// TIA Portal project "V1.0Final" (V17)

(* hardware
DEVICE "S7-1200 station_1"  S7-1200 Station
   slot 0: "Rack_0"  S7-1200 Rack  Rack  V1.0
   slot 1: "PLC_1"  CPU 1212C AC/DC/Rly  6ES7 212-1BD30-0XB0  V2.0
   slot 2: "AI 4x13BIT_1"  6ES7 231-4HD32-0XB0  V2.1
   slot 3: "AQ 2x14BIT_1"  SM 1232 AQ2  6ES7 232-4HB32-0XB0  V2.1
DEVICE "HMI_1"  KTP700 Basic PN
   slot 0: "HMI_1"  KTP700 Basic PN  6AV2 123-2GB03-0AX0  17.0.0.0
   slot 1: "HMI_RT_1"  KTP700 Basic PN  6AV2 123-2GB03-0AX0  17.0.0.0
   slot 5: "HMI_1.IE_CP_1"  PROFINET Interface  17.0.0.0
      slot 1: "PROFINET Interface_1"  PROFINET Interface
         slot 1: "Port_1"  Port
*)

// ===== PLC "PLC_1"  CPU 1212C AC/DC/Rly =====

VAR_GLOBAL   // PLC tag table "Default tag table"
   "DI_EM_STOP" AT %I0.0 : Bool;
   "DI_LS_Tørrkjøringsvern" AT %I0.1 : Bool;
   "DI_Reset_EM_STOP" AT %I0.2 : Bool;
   "AI_LT_01" AT %IW100 : Int;
   "DQ_Lys_EM_STOP" AT %Q0.1 : Bool;
   "AQ1_PÅDRAG_PUMPE_01" AT %QW112 : Int;
   "AQ2" AT %QW114 : Int;
   "DI_PUMPE_01_KJØRER" AT %I0.3 : Bool;
   "Tag_1" AT %M0.0 : Bool;
   "DQ_START_PUMPE_01" AT %Q0.2 : Bool;
   "AI_Hastighet_P01" AT %IW102 : Int;
END_VAR

// folder: Equipment

TYPE "UDT_Analog_Konvertering"
   STRUCT
      CFG : Struct   // Configuration Data
         Spare : Bool;
      END_STRUCT;
      Sts : Struct   // Status Data
         EU_Verdi_Out : Real;
      END_STRUCT;
      Cmd : Struct   // Command and request Data
         Spare : Bool;
      END_STRUCT;
      Par : Struct   // Parameter Data
         EU_Min : Real;
         EU_Max : Real;
      END_STRUCT;
      Fit : Struct   // Warning and alarm triggers
         Feil : Bool;
      END_STRUCT;
      Spare : Bool;   // False
   END_STRUCT;
END_TYPE

TYPE "UDT_Pumpe_Kontroll"
   STRUCT
      CFG : Struct
         Spare : Bool;
      END_STRUCT;
      Sts : Struct
         Pumpe_Run : Bool;
         Pumpe_Status : Int;
         Pumpe_Faktisk_Hastighet_Fra_VFD : Real;
         Pumpe_Pådrag_Fra_PID_Blokk : Real;
      END_STRUCT;
      Cmd : Struct
         Man_Start_Pumpe : Bool;
         Man_Stop_Pumpe : Bool;
         Auto_Start_Pumpe : Bool;
         EM_Stop : Bool;
         Tørrkjøringsvakt_LS_01 : Bool;
      END_STRUCT;
      Par : Struct
         Pådrag_Fra_PID_Blokk : Int;
      END_STRUCT;
      Fit : Struct
         Feil : Bool;
      END_STRUCT;
   END_STRUCT;
END_TYPE

// folder: Machine

TYPE "UDT_HMI"
   STRUCT
      CFG : Struct
         Spare : Bool;
      END_STRUCT;
      Sts : Struct
         HMI_PV : Real;
         HMI_Pump_Status : Int;
      END_STRUCT;
      Cmd : Struct
         HMI_Pump_Auto : Bool;
         HMI_Pump_Manuell : Bool;
         HMI_Pump_Start : Bool;
         HMI_Pump_Stop : Bool;
         HMI_Reset_Alarm : Bool;
         Spare : Bool;
      END_STRUCT;
      Par : Struct
         HMI_P_Gain : Real;
         HMI_Ti : Real;
         HMI_Td : Real;
         HMI_Manual_Speed_Ref : Real;
         HMI_LT_Level_SP : Real;
         HMI_LT_EU_Min : Real;
         HMI_LT_EU_Max : Real;
         HMI_Anti_Windup : Bool;
         Spare : Bool;
      END_STRUCT;
      Fit : Struct
         HMI_EM_Stop_Alarm : Bool;
         HMI_LS_Activated : Bool;
         HMI_Fault_Timer_SP : Time;
         HMI_Fault : Bool;
      END_STRUCT;
   END_STRUCT;
END_TYPE

// folder: (top level)

DATA_BLOCK "LT_01"   // DB6
{ S7_Optimized_Access := 'TRUE' }
VERSION : 0.1
// stored: InstanceOfName Analog_Konvertering
"Analog_Konvertering"
BEGIN
END_DATA_BLOCK

DATA_BLOCK "Pumpe_01_Kontroll_DB"   // DB8
{ S7_Optimized_Access := 'TRUE' }
VERSION : 0.1
// stored: InstanceOfName Pumpe_Kontroll
"Pumpe_Kontroll"
BEGIN
END_DATA_BLOCK

DATA_BLOCK "Regulerings_Rig_01_DB"   // DB9
{ S7_Optimized_Access := 'TRUE' }
VERSION : 0.1
// stored: InstanceOfName Regulerings_Rig
"Regulerings_Rig"
BEGIN
END_DATA_BLOCK

DATA_BLOCK "VFD_AQ_Hastighet_Pumpe01_DB"   // DB11
{ S7_Optimized_Access := 'TRUE' }
VERSION : 0.1
// stored: InstanceOfName Analog_Konvertering
"Analog_Konvertering"
BEGIN
END_DATA_BLOCK

// folder: Global_Data

DATA_BLOCK "DB_Equipment"   // DB3
{ S7_Optimized_Access := 'TRUE' }
VERSION : 0.1
   VAR
      Pumpe_01_Kontroll : "UDT_Pumpe_Kontroll";
   END_VAR
   VAR RETAIN
      LT_01_Kontrolll : "UDT_Analog_Konvertering";
      HMI_Kontroll_Pumpe_01 : "UDT_HMI";
   END_VAR
   VAR
      VFD_01_Speed : "UDT_Analog_Konvertering";
   END_VAR
BEGIN
END_DATA_BLOCK

DATA_BLOCK "DB_Machine"   // DB4
{ S7_Optimized_Access := 'TRUE' }
VERSION : 0.1
   VAR
      HMI_Control : "UDT_HMI";
   END_VAR
BEGIN
END_DATA_BLOCK

// folder: System blocks/Program resources

DATA_BLOCK "EM_Stop_TON_DB"   // DB1
{ S7_Optimized_Access := 'TRUE' }
AUTHOR : Simatic
FAMILY : IEC
NAME : IEC_TMR
VERSION : 1.0
// stored: InstanceOfName IEC_TIMER
"IEC_TIMER"
BEGIN
END_DATA_BLOCK

DATA_BLOCK "EM_Stop_TOF_DB"   // DB2
{ S7_Optimized_Access := 'TRUE' }
AUTHOR : Simatic
FAMILY : IEC
NAME : IEC_TMR
VERSION : 1.0
// stored: InstanceOfName IEC_TIMER
"IEC_TIMER"
BEGIN
END_DATA_BLOCK

DATA_BLOCK "Pump_Fault_Timer_DB"   // DB5
{ S7_Optimized_Access := 'TRUE' }
AUTHOR : Simatic
FAMILY : IEC
NAME : IEC_TMR
VERSION : 1.0
// stored: InstanceOfName IEC_TIMER
"IEC_TIMER"
BEGIN
END_DATA_BLOCK

// folder: (top level)

ORGANIZATION_BLOCK "Main"   // OB1, LAD, ProgramCycle
TITLE = "Main Program Sweep (Cycle)"
{ S7_Optimized_Access := 'TRUE' }
VERSION : 0.1
BEGIN
END_ORGANIZATION_BLOCK

ORGANIZATION_BLOCK "Cyclic interrupt"   // OB30, LAD, CyclicInterrupt
{ S7_Optimized_Access := 'TRUE' }
VERSION : 0.1
   VAR_TEMP
      "0" : Bool;
   END_VAR
BEGIN

REGION Network 1
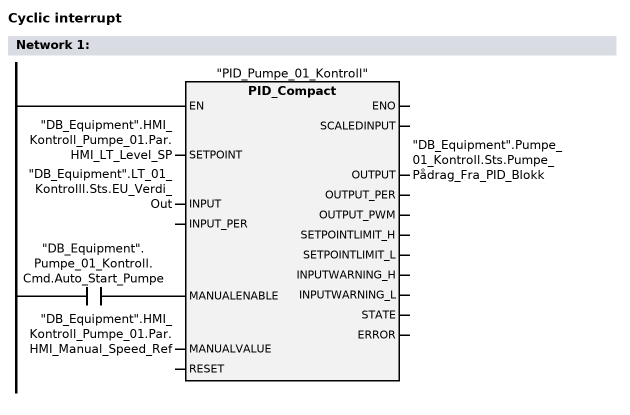
   "PID_Pumpe_01_Kontroll"(Setpoint := "DB_Equipment".HMI_Kontroll_Pumpe_01.Par.HMI_LT_Level_SP,   // PID_Compact
                           Input := "DB_Equipment".LT_01_Kontrolll.Sts.EU_Verdi_Out,
                           ManualEnable := "DB_Equipment".Pumpe_01_Kontroll.Cmd.Auto_Start_Pumpe,
                           ManualValue := "DB_Equipment".HMI_Kontroll_Pumpe_01.Par.HMI_Manual_Speed_Ref,
                           Output => "DB_Equipment".Pumpe_01_Kontroll.Sts.Pumpe_Pådrag_Fra_PID_Blokk);
END_REGION
END_ORGANIZATION_BLOCK

ORGANIZATION_BLOCK "Machine"   // OB123, LAD, ProgramCycle
TITLE = "Main Program Sweep (Cycle)"
{ S7_Optimized_Access := 'TRUE' }
VERSION : 0.1
BEGIN

REGION Network 1
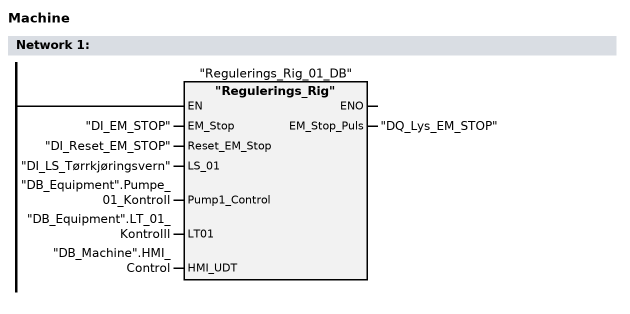
   RUNG wire#powerrail
      "Regulerings_Rig_01_DB"(EM_Stop := "DI_EM_STOP", Reset_EM_Stop := "DI_Reset_EM_STOP", LS_01 := "DI_LS_Tørrkjøringsvern", Pump1_Control := "DB_Equipment".Pumpe_01_Kontroll, LT01 := "DB_Equipment".LT_01_Kontrolll, HMI_UDT := "DB_Machine".HMI_Control, EM_Stop_Puls => "DQ_Lys_EM_STOP")
   END_RUNG
   // the same network as SCL:
   "Regulerings_Rig_01_DB"(EM_Stop := "DI_EM_STOP",   // "Regulerings_Rig"
                           Reset_EM_Stop := "DI_Reset_EM_STOP",
                           LS_01 := "DI_LS_Tørrkjøringsvern",
                           Pump1_Control := "DB_Equipment".Pumpe_01_Kontroll,
                           LT01 := "DB_Equipment".LT_01_Kontrolll,
                           HMI_UDT := "DB_Machine".HMI_Control,
                           EM_Stop_Puls => "DQ_Lys_EM_STOP");
END_REGION
END_ORGANIZATION_BLOCK

ORGANIZATION_BLOCK "Equipment"   // OB124, LAD, ProgramCycle
TITLE = "Main Program Sweep (Cycle)"
{ S7_Optimized_Access := 'TRUE' }
VERSION : 0.1
BEGIN

REGION Network 1
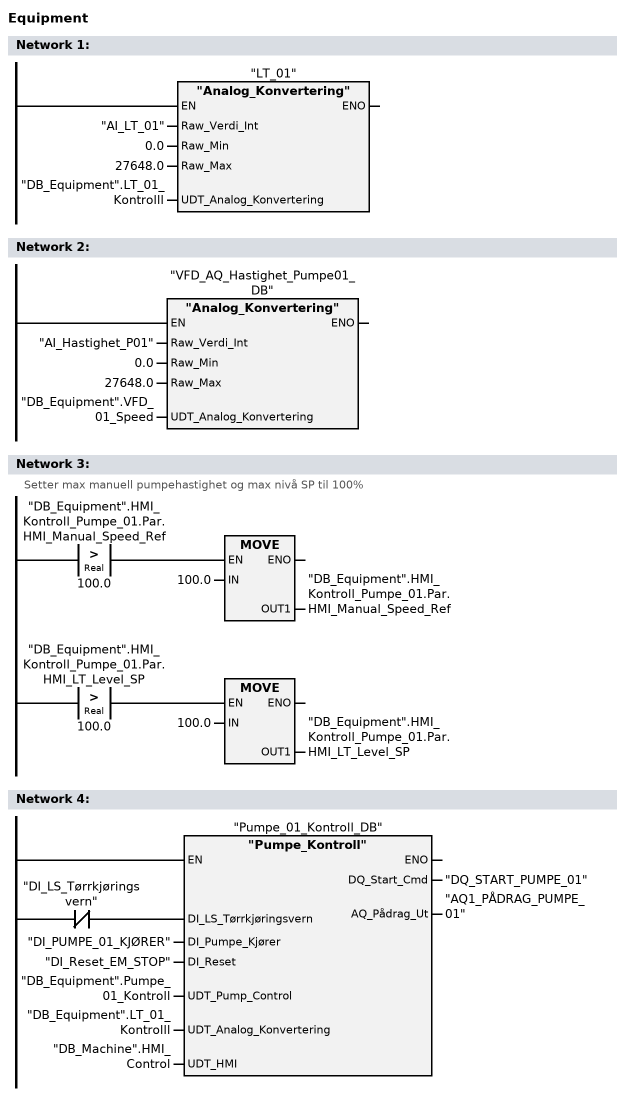
   RUNG wire#powerrail
      "LT_01"(Raw_Verdi_Int := "AI_LT_01", Raw_Min := 0.0, Raw_Max := 27648.0, UDT_Analog_Konvertering := "DB_Equipment".LT_01_Kontrolll)
   END_RUNG
   // the same network as SCL:
   "LT_01"(Raw_Verdi_Int := "AI_LT_01",   // "Analog_Konvertering"
           Raw_Min := 0.0,
           Raw_Max := 27648.0,
           UDT_Analog_Konvertering := "DB_Equipment".LT_01_Kontrolll);
END_REGION

REGION Network 2
   RUNG wire#powerrail
      "VFD_AQ_Hastighet_Pumpe01_DB"(Raw_Verdi_Int := "AI_Hastighet_P01", Raw_Min := 0.0, Raw_Max := 27648.0, UDT_Analog_Konvertering := "DB_Equipment".VFD_01_Speed)
   END_RUNG
   // the same network as SCL:
   "VFD_AQ_Hastighet_Pumpe01_DB"(Raw_Verdi_Int := "AI_Hastighet_P01",   // "Analog_Konvertering"
                           Raw_Min := 0.0,
                           Raw_Max := 27648.0,
                           UDT_Analog_Konvertering := "DB_Equipment".VFD_01_Speed);
END_REGION

REGION Network 3
   // Setter max manuell pumpehastighet og max nivå SP til 100%
   RUNG wire#powerrail
      { S7_Templates := "SrcType := Real" } GT_Contact(in1 := "DB_Equipment".HMI_Kontroll_Pumpe_01.Par.HMI_Manual_Speed_Ref, in2 := 100.0)
      { S7_GenerateENO := "TRUE" } Move(in := 100.0, out1 => "DB_Equipment".HMI_Kontroll_Pumpe_01.Par.HMI_Manual_Speed_Ref)
   END_RUNG
   RUNG wire#powerrail
      { S7_Templates := "SrcType := Real" } GT_Contact(in1 := "DB_Equipment".HMI_Kontroll_Pumpe_01.Par.HMI_LT_Level_SP, in2 := 100.0)
      { S7_GenerateENO := "TRUE" } Move(in := 100.0, out1 => "DB_Equipment".HMI_Kontroll_Pumpe_01.Par.HMI_LT_Level_SP)
   END_RUNG
   // the same network as SCL:
   IF "DB_Equipment".HMI_Kontroll_Pumpe_01.Par.HMI_Manual_Speed_Ref > 100.0 THEN
       "DB_Equipment".HMI_Kontroll_Pumpe_01.Par.HMI_Manual_Speed_Ref := 100.0;
   END_IF;
   IF "DB_Equipment".HMI_Kontroll_Pumpe_01.Par.HMI_LT_Level_SP > 100.0 THEN
       "DB_Equipment".HMI_Kontroll_Pumpe_01.Par.HMI_LT_Level_SP := 100.0;
   END_IF;
END_REGION

REGION Network 4
   RUNG wire#powerrail
      "Pumpe_01_Kontroll_DB"(DI_LS_Tørrkjøringsvern := wire#w1, DI_Pumpe_Kjører := "DI_PUMPE_01_KJØRER", DI_Reset := "DI_Reset_EM_STOP", UDT_Pump_Control := "DB_Equipment".Pumpe_01_Kontroll, UDT_Analog_Konvertering := "DB_Equipment".LT_01_Kontrolll, UDT_HMI := "DB_Machine".HMI_Control, DQ_Start_Cmd => "DQ_START_PUMPE_01", AQ_Pådrag_Ut => "AQ1_PÅDRAG_PUMPE_01")
   END_RUNG
   RUNG wire#powerrail
      I_Contact( "DI_LS_Tørrkjøringsvern" )
   END_RUNG wire#w1
   // the same network as SCL:
   "Pumpe_01_Kontroll_DB"(DI_LS_Tørrkjøringsvern := NOT "DI_LS_Tørrkjøringsvern",   // "Pumpe_Kontroll"
                          DI_Pumpe_Kjører := "DI_PUMPE_01_KJØRER",
                          DI_Reset := "DI_Reset_EM_STOP",
                          UDT_Pump_Control := "DB_Equipment".Pumpe_01_Kontroll,
                          UDT_Analog_Konvertering := "DB_Equipment".LT_01_Kontrolll,
                          UDT_HMI := "DB_Machine".HMI_Control,
                          DQ_Start_Cmd => "DQ_START_PUMPE_01",
                          AQ_Pådrag_Ut => "AQ1_PÅDRAG_PUMPE_01");
END_REGION
END_ORGANIZATION_BLOCK

// folder: Equipment

FUNCTION_BLOCK "Analog_Konvertering"   // FB2, LAD
{ S7_Optimized_Access := 'TRUE' }
VERSION : 0.1
   VAR_INPUT
      Raw_Verdi_Int : Int;
      Raw_Min : Real;
      Raw_Max : Real;
   END_VAR
   VAR_IN_OUT
      UDT_Analog_Konvertering : "UDT_Analog_Konvertering";
   END_VAR
   VAR
      Convert_Value : Real;
      Raw_Value_Real : Real;
      EU_Value_Real : Real;
   END_VAR
BEGIN

REGION Network 1
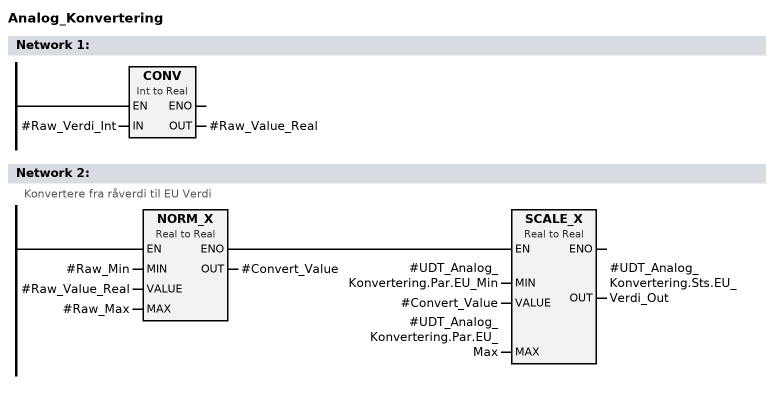
   RUNG wire#powerrail
      { S7_Templates := "[SrcType := Int, DestType := Real]"; S7_GenerateENO := "TRUE" } Convert(in := #Raw_Verdi_Int, out => #Raw_Value_Real)
   END_RUNG
   // the same network as SCL:
   #Raw_Value_Real := INT_TO_REAL(#Raw_Verdi_Int);
END_REGION

REGION Network 2
   // Konvertere fra råverdi til EU Verdi
   RUNG wire#powerrail
      { S7_Templates := "[SrcType := Real, DestType := Real]"; S7_GenerateENO := "TRUE" } Normalize(min := #Raw_Min, value := #Raw_Value_Real, max := #Raw_Max, out => #Convert_Value)
      { S7_Templates := "[SrcType := Real, DestType := Real]"; S7_GenerateENO := "TRUE" } Scale(min := #UDT_Analog_Konvertering.Par.EU_Min, value := #Convert_Value, max := #UDT_Analog_Konvertering.Par.EU_Max, out => #UDT_Analog_Konvertering.Sts.EU_Verdi_Out)
   END_RUNG
   // the same network as SCL:
   // ENO of a box is taken as its EN; it also drops when the box reports an error
   #Convert_Value := NORM_X(MIN := #Raw_Min, VALUE := #Raw_Value_Real, MAX := #Raw_Max);
   #UDT_Analog_Konvertering.Sts.EU_Verdi_Out := SCALE_X(MIN := #UDT_Analog_Konvertering.Par.EU_Min, VALUE := #Convert_Value, MAX := #UDT_Analog_Konvertering.Par.EU_Max);
END_REGION
END_FUNCTION_BLOCK

FUNCTION_BLOCK "Pumpe_Kontroll"   // FB3, LAD
{ S7_Optimized_Access := 'TRUE' }
VERSION : 0.1
   VAR_INPUT
      DI_LS_Tørrkjøringsvern : Bool;
      DI_Pumpe_Kjører : Bool;
      DI_Reset : Bool;
   END_VAR
   VAR_OUTPUT
      DQ_Start_Cmd : Bool;
      AQ_Pådrag_Ut : Int;
   END_VAR
   VAR_IN_OUT
      UDT_Pump_Control : "UDT_Pumpe_Kontroll";
      UDT_Analog_Konvertering : "UDT_Analog_Konvertering";
      UDT_HMI : "UDT_HMI";
   END_VAR
   VAR
      Tmp_Start_Cmd_Man : Bool;
      Tmp_Start_Cmd_Auto : Bool;
      Tmp_Pådrag_Ut_Int : Int;
      Tmp_Pådrag_Ut_Real : Real;
      Convert_Value : Real;
   END_VAR
BEGIN

REGION Network 1
   // Manuell Start og stopp kriterier
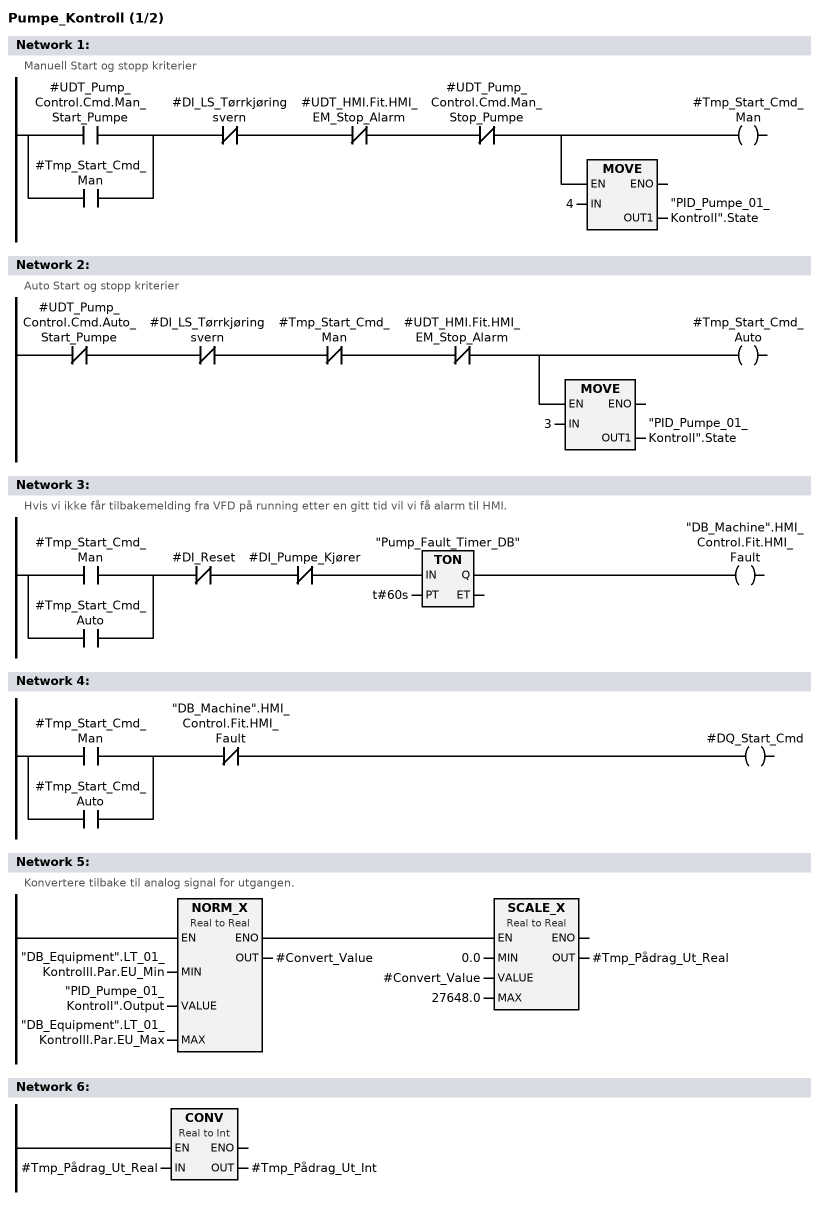
   RUNG wire#powerrail
      Contact( #UDT_Pump_Control.Cmd.Man_Start_Pumpe )
      wire#w1
      I_Contact( #DI_LS_Tørrkjøringsvern )
      I_Contact( #UDT_HMI.Fit.HMI_EM_Stop_Alarm )
      I_Contact( #UDT_Pump_Control.Cmd.Man_Stop_Pumpe )
      wire#w2
      Coil( #Tmp_Start_Cmd_Man )
   END_RUNG
   RUNG wire#powerrail
      Contact( #Tmp_Start_Cmd_Man )
   END_RUNG wire#w1
   RUNG wire#w2
      { S7_GenerateENO := "TRUE" } Move(in := 4, out1 => "PID_Pumpe_01_Kontroll".State)
   END_RUNG
   // the same network as SCL:
   #Tmp_Start_Cmd_Man := (#UDT_Pump_Control.Cmd.Man_Start_Pumpe OR #Tmp_Start_Cmd_Man) AND NOT #DI_LS_Tørrkjøringsvern AND NOT #UDT_HMI.Fit.HMI_EM_Stop_Alarm AND NOT #UDT_Pump_Control.Cmd.Man_Stop_Pumpe;
   IF #Tmp_Start_Cmd_Man THEN "PID_Pumpe_01_Kontroll".State := 4; END_IF;
END_REGION

REGION Network 2
   // Auto Start og stopp kriterier
   RUNG wire#powerrail
      I_Contact( #UDT_Pump_Control.Cmd.Auto_Start_Pumpe )
      I_Contact( #DI_LS_Tørrkjøringsvern )
      I_Contact( #Tmp_Start_Cmd_Man )
      I_Contact( #UDT_HMI.Fit.HMI_EM_Stop_Alarm )
      wire#w1
      Coil( #Tmp_Start_Cmd_Auto )
   END_RUNG
   RUNG wire#w1
      { S7_GenerateENO := "TRUE" } Move(in := 3, out1 => "PID_Pumpe_01_Kontroll".State)
   END_RUNG
   // the same network as SCL:
   #Tmp_Start_Cmd_Auto := NOT #UDT_Pump_Control.Cmd.Auto_Start_Pumpe AND NOT #DI_LS_Tørrkjøringsvern AND NOT #Tmp_Start_Cmd_Man AND NOT #UDT_HMI.Fit.HMI_EM_Stop_Alarm;
   IF #Tmp_Start_Cmd_Auto THEN "PID_Pumpe_01_Kontroll".State := 3; END_IF;
END_REGION

REGION Network 3
   // Hvis vi ikke får tilbakemelding fra VFD på running etter en gitt tid vil vi få alarm til HMI.
   "Pump_Fault_Timer_DB".TON(IN := (#Tmp_Start_Cmd_Man OR #Tmp_Start_Cmd_Auto) AND NOT #DI_Reset AND NOT #DI_Pumpe_Kjører,
                           PT := t#60s);
   "DB_Machine".HMI_Control.Fit.HMI_Fault := "Pump_Fault_Timer_DB".Q;
END_REGION

REGION Network 4
   RUNG wire#powerrail
      Contact( #Tmp_Start_Cmd_Man )
      wire#w1
      I_Contact( "DB_Machine".HMI_Control.Fit.HMI_Fault )
      Coil( #DQ_Start_Cmd )
   END_RUNG
   RUNG wire#powerrail
      Contact( #Tmp_Start_Cmd_Auto )
   END_RUNG wire#w1
   // the same network as SCL:
   #DQ_Start_Cmd := (#Tmp_Start_Cmd_Man OR #Tmp_Start_Cmd_Auto) AND NOT "DB_Machine".HMI_Control.Fit.HMI_Fault;
END_REGION

REGION Network 5
   // Konvertere tilbake til analog signal for utgangen.
   RUNG wire#powerrail
      { S7_Templates := "[SrcType := Real, DestType := Real]"; S7_GenerateENO := "TRUE" } Normalize(min := "DB_Equipment".LT_01_Kontrolll.Par.EU_Min, value := "PID_Pumpe_01_Kontroll".Output, max := "DB_Equipment".LT_01_Kontrolll.Par.EU_Max, out => #Convert_Value)
      { S7_Templates := "[SrcType := Real, DestType := Real]"; S7_GenerateENO := "TRUE" } Scale(min := 0.0, value := #Convert_Value, max := 27648.0, out => #Tmp_Pådrag_Ut_Real)
   END_RUNG
   // the same network as SCL:
   // ENO of a box is taken as its EN; it also drops when the box reports an error
   #Convert_Value := NORM_X(MIN := "DB_Equipment".LT_01_Kontrolll.Par.EU_Min, VALUE := "PID_Pumpe_01_Kontroll".Output, MAX := "DB_Equipment".LT_01_Kontrolll.Par.EU_Max);
   #Tmp_Pådrag_Ut_Real := SCALE_X(MIN := 0.0, VALUE := #Convert_Value, MAX := 27648.0);
END_REGION

REGION Network 6
   RUNG wire#powerrail
      { S7_Templates := "[SrcType := Real, DestType := Int]"; S7_GenerateENO := "TRUE" } Convert(in := #Tmp_Pådrag_Ut_Real, out => #Tmp_Pådrag_Ut_Int)
   END_RUNG
   // the same network as SCL:
   #Tmp_Pådrag_Ut_Int := REAL_TO_INT(#Tmp_Pådrag_Ut_Real);
END_REGION

REGION Network 7
   // Når vi har start signal vil pådraget overføres fra PID blokk til Analog utgang for pådrag til pumpe.
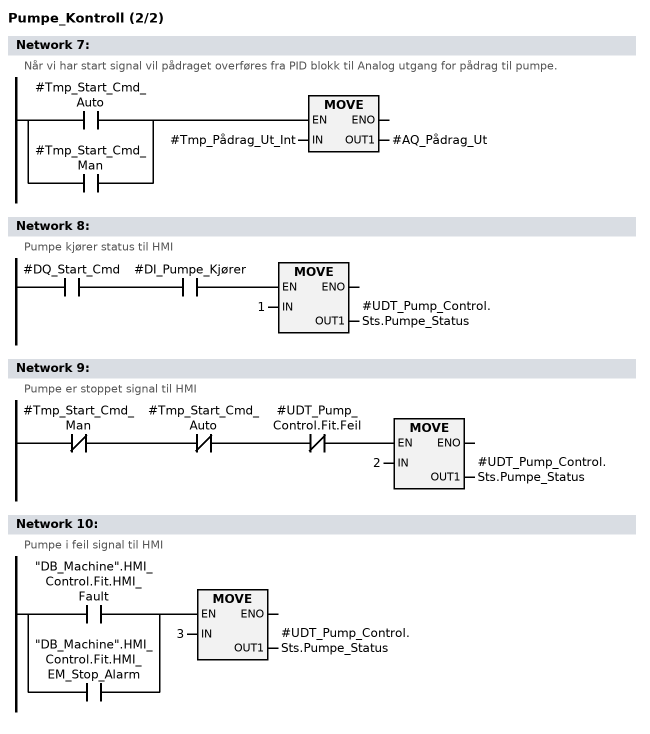
   RUNG wire#powerrail
      Contact( #Tmp_Start_Cmd_Auto )
      wire#w1
      { S7_GenerateENO := "TRUE" } Move(in := #Tmp_Pådrag_Ut_Int, out1 => #AQ_Pådrag_Ut)
   END_RUNG
   RUNG wire#powerrail
      Contact( #Tmp_Start_Cmd_Man )
   END_RUNG wire#w1
   // the same network as SCL:
   IF #Tmp_Start_Cmd_Auto OR #Tmp_Start_Cmd_Man THEN #AQ_Pådrag_Ut := #Tmp_Pådrag_Ut_Int; END_IF;
END_REGION

REGION Network 8
   // Pumpe kjører status til HMI
   RUNG wire#powerrail
      Contact( #DQ_Start_Cmd )
      Contact( #DI_Pumpe_Kjører )
      { S7_GenerateENO := "TRUE" } Move(in := 1, out1 => #UDT_Pump_Control.Sts.Pumpe_Status)
   END_RUNG
   // the same network as SCL:
   IF #DQ_Start_Cmd AND #DI_Pumpe_Kjører THEN #UDT_Pump_Control.Sts.Pumpe_Status := 1; END_IF;
END_REGION

REGION Network 9
   // Pumpe er stoppet signal til HMI
   RUNG wire#powerrail
      I_Contact( #Tmp_Start_Cmd_Man )
      I_Contact( #Tmp_Start_Cmd_Auto )
      I_Contact( #UDT_Pump_Control.Fit.Feil )
      { S7_GenerateENO := "TRUE" } Move(in := 2, out1 => #UDT_Pump_Control.Sts.Pumpe_Status)
   END_RUNG
   // the same network as SCL:
   IF NOT #Tmp_Start_Cmd_Man AND NOT #Tmp_Start_Cmd_Auto AND NOT #UDT_Pump_Control.Fit.Feil THEN
       #UDT_Pump_Control.Sts.Pumpe_Status := 2;
   END_IF;
END_REGION

REGION Network 10
   // Pumpe i feil signal til HMI
   RUNG wire#powerrail
      Contact( "DB_Machine".HMI_Control.Fit.HMI_Fault )
      wire#w1
      { S7_GenerateENO := "TRUE" } Move(in := 3, out1 => #UDT_Pump_Control.Sts.Pumpe_Status)
   END_RUNG
   RUNG wire#powerrail
      Contact( "DB_Machine".HMI_Control.Fit.HMI_EM_Stop_Alarm )
   END_RUNG wire#w1
   // the same network as SCL:
   IF "DB_Machine".HMI_Control.Fit.HMI_Fault OR "DB_Machine".HMI_Control.Fit.HMI_EM_Stop_Alarm THEN
       #UDT_Pump_Control.Sts.Pumpe_Status := 3;
   END_IF;
END_REGION
END_FUNCTION_BLOCK

// folder: Machine

FUNCTION_BLOCK "Regulerings_Rig"   // FB1, LAD
{ S7_Optimized_Access := 'TRUE' }
VERSION : 0.1
   VAR_INPUT
      EM_Stop : Bool;
      Reset_EM_Stop : Bool;
      LS_01 : Bool;
   END_VAR
   VAR_OUTPUT
      EM_Stop_Puls : Bool;
   END_VAR
   VAR_IN_OUT
      Pump1_Control : "UDT_Pumpe_Kontroll";
      LT01 : "UDT_Analog_Konvertering";
      HMI_UDT : "UDT_HMI";
   END_VAR
   VAR
      Tmp_EM_Stop_Alarm : Bool;
      Tmp_Enable_PID : Bool;
      Tmp_Blink_Off : Bool;
      Tmp_Blink_On : Bool;
      Tmp_LS_Alarm : Bool;
   END_VAR
BEGIN

REGION Network 1
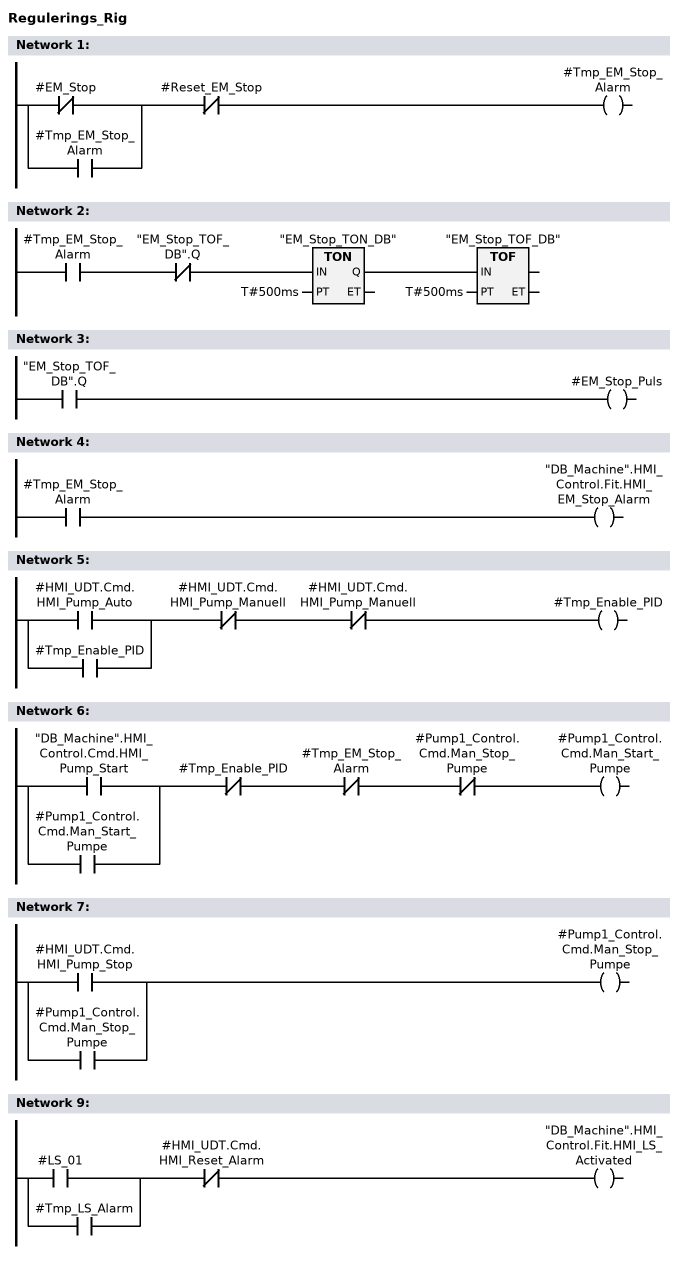
   RUNG wire#powerrail
      I_Contact( #EM_Stop )
      wire#w1
      I_Contact( #Reset_EM_Stop )
      Coil( #Tmp_EM_Stop_Alarm )
   END_RUNG
   RUNG wire#powerrail
      Contact( #Tmp_EM_Stop_Alarm )
   END_RUNG wire#w1
   // the same network as SCL:
   #Tmp_EM_Stop_Alarm := (NOT #EM_Stop OR #Tmp_EM_Stop_Alarm) AND NOT #Reset_EM_Stop;
END_REGION

REGION Network 2
   "EM_Stop_TON_DB".TON(IN := #Tmp_EM_Stop_Alarm AND NOT "EM_Stop_TOF_DB".Q, PT := T#500ms);
   "EM_Stop_TOF_DB".TOF(IN := "EM_Stop_TON_DB".Q, PT := T#500ms);
END_REGION

REGION Network 3
   RUNG wire#powerrail
      Contact( "EM_Stop_TOF_DB".Q )
      Coil( #EM_Stop_Puls )
   END_RUNG
   // the same network as SCL:
   #EM_Stop_Puls := "EM_Stop_TOF_DB".Q;
END_REGION

REGION Network 4
   RUNG wire#powerrail
      Contact( #Tmp_EM_Stop_Alarm )
      Coil( "DB_Machine".HMI_Control.Fit.HMI_EM_Stop_Alarm )
   END_RUNG
   // the same network as SCL:
   "DB_Machine".HMI_Control.Fit.HMI_EM_Stop_Alarm := #Tmp_EM_Stop_Alarm;
END_REGION

REGION Network 5
   RUNG wire#powerrail
      Contact( #HMI_UDT.Cmd.HMI_Pump_Auto )
      wire#w1
      I_Contact( #HMI_UDT.Cmd.HMI_Pump_Manuell )
      I_Contact( #HMI_UDT.Cmd.HMI_Pump_Manuell )
      Coil( #Tmp_Enable_PID )
   END_RUNG
   RUNG wire#powerrail
      Contact( #Tmp_Enable_PID )
   END_RUNG wire#w1
   // the same network as SCL:
   #Tmp_Enable_PID := (#HMI_UDT.Cmd.HMI_Pump_Auto OR #Tmp_Enable_PID) AND NOT #HMI_UDT.Cmd.HMI_Pump_Manuell AND NOT #HMI_UDT.Cmd.HMI_Pump_Manuell;
END_REGION

REGION Network 6
   RUNG wire#powerrail
      Contact( "DB_Machine".HMI_Control.Cmd.HMI_Pump_Start )
      wire#w1
      I_Contact( #Tmp_Enable_PID )
      I_Contact( #Tmp_EM_Stop_Alarm )
      I_Contact( #Pump1_Control.Cmd.Man_Stop_Pumpe )
      Coil( #Pump1_Control.Cmd.Man_Start_Pumpe )
   END_RUNG
   RUNG wire#powerrail
      Contact( #Pump1_Control.Cmd.Man_Start_Pumpe )
   END_RUNG wire#w1
   // the same network as SCL:
   #Pump1_Control.Cmd.Man_Start_Pumpe := ("DB_Machine".HMI_Control.Cmd.HMI_Pump_Start OR #Pump1_Control.Cmd.Man_Start_Pumpe) AND NOT #Tmp_Enable_PID AND NOT #Tmp_EM_Stop_Alarm AND NOT #Pump1_Control.Cmd.Man_Stop_Pumpe;
END_REGION

REGION Network 7
   RUNG wire#powerrail
      Contact( #HMI_UDT.Cmd.HMI_Pump_Stop )
      wire#w1
      Coil( #Pump1_Control.Cmd.Man_Stop_Pumpe )
   END_RUNG
   RUNG wire#powerrail
      Contact( #Pump1_Control.Cmd.Man_Stop_Pumpe )
   END_RUNG wire#w1
   // the same network as SCL:
   #Pump1_Control.Cmd.Man_Stop_Pumpe := #HMI_UDT.Cmd.HMI_Pump_Stop OR #Pump1_Control.Cmd.Man_Stop_Pumpe;
END_REGION

REGION Network 9
   RUNG wire#powerrail
      Contact( #LS_01 )
      wire#w1
      I_Contact( #HMI_UDT.Cmd.HMI_Reset_Alarm )
      Coil( "DB_Machine".HMI_Control.Fit.HMI_LS_Activated )
   END_RUNG
   RUNG wire#powerrail
      Contact( #Tmp_LS_Alarm )
   END_RUNG wire#w1
   // the same network as SCL:
   "DB_Machine".HMI_Control.Fit.HMI_LS_Activated := (#LS_01 OR #Tmp_LS_Alarm) AND NOT #HMI_UDT.Cmd.HMI_Reset_Alarm;
END_REGION
END_FUNCTION_BLOCK

(* ===== HMI "HMI_RT_1" =====
system functions are stored by id; their names below are inferred from use
connection "HMI_Connection_1": ETHERNET, SMART_S7_1200_OMS

HMI tags "Default tag table"
   "DB_Equipment_HMI_Control_Par_HMI_P_Gain" : Real = PLC DB_Equipment.HMI_Kontroll_Pumpe_01.Par.HMI_Ti, 1 s
   "DB_Equipment_HMI_Control_Pump1" : UDT_HMI = PLC DB_Equipment.HMI_Kontroll_Pumpe_01, 1 s
   "DB_Machine_HMI_Control_Par_HMI_Ti" : Real = PLC DB_Machine.HMI_Control.Par.HMI_Ti, 1 s
   "DB_Equipment_HMI_Control_Pump1_Par_HMI_P_Gain" : Real = PLC DB_Equipment.HMI_Kontroll_Pumpe_01.Par.HMI_P_Gain, 1 s
   "DB_Equipment_HMI_Control_Pump1_Par_HMI_Td" : Real = PLC DB_Equipment.HMI_Kontroll_Pumpe_01.Par.HMI_Td, 1 s
   "DB_Equipment_HMI_Control_Pump1_Sts_HMI_Level_PV" : Real = PLC DB_Equipment.HMI_Kontroll_Pumpe_01.Sts.HMI_PV, 1 s
   "LT_01_Raw_Min" : Real = PLC LT_01.Raw_Min, 1 s
   "LT_01_Raw_Max" : Real = PLC LT_01.Raw_Max, 1 s
   "DB_Equipment_HMI_Control_Pump1_Cmd_HMI_Pump_Manuell" : Bool = PLC DB_Equipment.HMI_Kontroll_Pumpe_01.Cmd.HMI_Pump_Manuell, 1 s
   "DB_Equipment_HMI_Control_Pump1_Cmd_HMI_Pump_Auto" : Bool = PLC DB_Equipment.HMI_Kontroll_Pumpe_01.Cmd.HMI_Pump_Auto, 1 s
   "DB_Equipment_HMI_Control_Pump1_Cmd_HMI_Pump_Start" : Bool = PLC DB_Equipment.HMI_Kontroll_Pumpe_01.Cmd.HMI_Pump_Start, 1 s
   "DB_Equipment_HMI_Control_Pump1_Cmd_HMI_Pump_Stop" : Bool = PLC DB_Equipment.HMI_Kontroll_Pumpe_01.Cmd.HMI_Pump_Stop, 1 s
   "DB_Equipment_HMI_Control_Pump1_Par_HMI_Manual_Speed_Ref" : Real = PLC DB_Equipment.HMI_Kontroll_Pumpe_01.Par.HMI_Manual_Speed_Ref, 1 s
   "DB_Machine_HMI_Control_Sts_HMI_PV" : Real = PLC DB_Machine.HMI_Control.Sts.HMI_PV, 1 s
   "DB_Equipment_LT01_Control_Sts_EU_Value_Out" : Real = PLC DB_Equipment.LT_01_Kontrolll.Sts.EU_Verdi_Out, 1 s
   "DB_Equipment_LT01_Control_Par_EU_Min" : Real = PLC DB_Equipment.LT_01_Kontrolll.Par.EU_Min, 1 s
   "DB_Equipment_LT01_Control_Par_EU_Max" : Real = PLC DB_Equipment.LT_01_Kontrolll.Par.EU_Max, 1 s
   "PID_Pump1_Control_sRet_r_Ctrl_Gain" : Real = PLC PID_Pumpe_01_Kontroll.sRet.r_Ctrl_Gain, 1 s
   "PID_Pump1_Control_sRet_r_Ctrl_Ti" : Real = PLC PID_Pumpe_01_Kontroll.sRet.r_Ctrl_Ti, 1 s
   "PID_Pump1_Control_sRet_r_Ctrl_Td" : Real = PLC PID_Pumpe_01_Kontroll.sRet.r_Ctrl_Td, 1 s
   "DI_P01_Run" : Bool = PLC DI_PUMPE_01_KJØRER AT %I0.3, 1 s
   "DB_Equipment_Pump1_Control_Sts_Pump_Aktuell_Hastighet" : Real = PLC DB_Equipment.Pumpe_01_Kontroll.Sts.Pumpe_Faktisk_Hastighet_Fra_VFD, 1 s
   "DB_Equipment_Pump1_Control_Sts_Pumpe_Pådrag_Fra_PID_Blokk" : Real = PLC DB_Equipment.Pumpe_01_Kontroll.Sts.Pumpe_Pådrag_Fra_PID_Blokk, 1 s
   "DB_Equipment_Pumpe_01_Kontroll_Sts_Pumpe_Status" : Int = PLC DB_Equipment.Pumpe_01_Kontroll.Sts.Pumpe_Status, 1 s
   "DB_Equipment_Pumpe_01_Kontroll_Cmd_Man_Start_Pumpe" : Bool = PLC DB_Equipment.Pumpe_01_Kontroll.Cmd.Man_Start_Pumpe, 1 s
   "DB_Equipment_Pumpe_01_Kontroll_Cmd_Man_Stop_Pumpe" : Bool = PLC DB_Equipment.Pumpe_01_Kontroll.Cmd.Man_Stop_Pumpe, 1 s
   "PID_Pumpe_01_Kontroll_sPid_Cmpt_r_Pv_Norm_OUT_1" : Real = PLC PID_Pumpe_01_Kontroll.sPid_Cmpt.r_Pv_Norm_OUT_1, 1 s
   "PID_Pumpe_01_Kontroll_Output" : Real = PLC PID_Pumpe_01_Kontroll.Output, 1 s
   "DB_Equipment_VFD_01_Speed_Sts_EU_Verdi_Out" : Real = PLC DB_Equipment.VFD_01_Speed.Sts.EU_Verdi_Out, 1 s
   "DB_Equipment_Pumpe_01_Kontroll_Cmd_Tørrkjøringsvakt_LS_01" : Bool = PLC DB_Equipment.Pumpe_01_Kontroll.Cmd.Tørrkjøringsvakt_LS_01, 1 s
   "DB_Machine_HMI_Control_Fit_HMI_LS_Activated" : Bool = PLC DB_Machine.HMI_Control.Fit.HMI_LS_Activated, 1 s
   "DB_Equipment_Pumpe_01_Kontroll_Cmd_Auto_Start_Pumpe" : Bool = PLC DB_Equipment.Pumpe_01_Kontroll.Cmd.Auto_Start_Pumpe, 1 s

screen "Prosess_Side" 800x480
   TextField "Text field_1" at 230,5 size 329x43; Text 'Team Level Legends'
   Bar "Bar_1" at 130,10 size 100x200; MinimumValue 0; MaximumValue 100
      ProcessValue <- "DB_Equipment_LT01_Control_Sts_EU_Value_Out"
   GraphicView "Graphic view_4" at 415,410 size 26x24; Picture "Graphic_7"
   GraphicView "Graphic view_5" at 172,392 size 197x25; Picture "Graphic_7"
   GraphicView "Graphic view_8" at 145,210 size 25x184; Picture "Graphic_9"
   GraphicView "Graphic view_9" at 195,210 size 25x25; Picture "Graphic_9"
   GraphicView "Graphic view_7" at 143,388 size 30x30; Picture "Graphic_10"
   GraphicView "Graphic view_2" at 197,232 size 25x45; Picture "Graphic_11"
   GraphicView "Graphic view_6" at 193,274 size 30x30; Picture "Graphic_10"
   GraphicView "Graphic view_10" at 222,277 size 291x25; Picture "Graphic_7"
   GraphicView "Graphic view_11" at 511,277 size 25x25; Picture "Graphic_12"
   GraphicView "Graphic view_12" at 511,299 size 25x52; Picture "Graphic_9"
   TextField "Text field_8" at 24,430 size 52x23; Text 'Setup'
   TextField "Text field_9" at 125,430 size 53x23; Text 'Trend'
   TextField "Text field_10" at 225,430 size 54x23; Text 'Alarm'
   TextField "Text field_16" at 29,450 size 40x23; Text 'Side'
   TextField "Text field_17" at 132,450 size 40x23; Text 'Side'
   TextField "Text field_18" at 230,450 size 40x23; Text 'Side'
   TextField "Text field_7" at 375,50 size 335x34; Text 'Pumpe 01 Manuell kjøring'
   TextField "Text field_11" at 360,100 size 336x34; Text 'Manuelt Pådrag Pumpe 01'
   IOField "I/O field_9" at 699,100 size 90x40; FormatPattern s999.9
      ProcessValue <- "DB_Equipment_HMI_Control_Pump1_Par_HMI_Manual_Speed_Ref"
   TextField "Text field_14" at 465,150 size 200x34; Text 'Start Pumpe 01'
   TextField "Text field_15" at 465,200 size 211x34; Text 'Stopp Pumpe 01'
   Button "Button_4" at 695,150 size 96x32; TextOff 'Start'
      on Press: function_b14e0dd5("DB_Equipment_Pumpe_01_Kontroll_Cmd_Man_Start_Pumpe", 0)
   Button "Button_5" at 693,200 size 96x32; TextOff 'Stopp'
      on Press: function_b14e0dd5("DB_Equipment_Pumpe_01_Kontroll_Cmd_Man_Stop_Pumpe", 0)
   TextField "Text field_2" at 241,304 size 260x34; Text 'Hastighet Pumpe 01'
   IOField "I/O field_1" at 345,344 size 90x40; FormatPattern s999.9
      ProcessValue <- "DB_Equipment_Pump1_Control_Sts_Pumpe_Pådrag_Fra_PID_Blokk"
   IOField "I/O field_2" at 20,105 size 90x40; FormatPattern s999.9
      ProcessValue <- "DB_Equipment_LT01_Control_Sts_EU_Value_Out"
   TextField "Text field_3" at 32,10 size 68x34; Text 'Nivå'
   TextField "Text field_4" at 5,40 size 124x34; Text 'Forbruks'
   TextField "Text field_5" at 32,70 size 66x34; Text 'Tank'
   Switch "Switch_1" at 726,50 size 64x32; TextOn 'ON'; CaptionText 'Switch'; TextOff 'OFF'
      ProcessValue <- "DB_Equipment_Pumpe_01_Kontroll_Cmd_Auto_Start_Pumpe"
   Circle "Circle_1" at 640,382 size 60x60
      Appearance <- "DB_Machine_HMI_Control_Fit_HMI_LS_Activated"
   TextField "Text field_6" at 648,400 size 44x23; Text 'LS01'
   Circle "Circle_2" at 365,380 size 60x60
      Appearance <- "DB_Equipment_Pumpe_01_Kontroll_Sts_Pumpe_Status"
   TextField "Text field_12" at 377,397 size 36x23; Text 'P01'
   Softkey "Softkey_F1" at 0,0 size 0x0
      on KeyDown: ActivateScreen("Setup_Side", 0)
   Softkey "Softkey_F2" at 0,0 size 0x0
      on KeyDown: ActivateScreen("Trend_Side", 0)
   Softkey "Softkey_F3" at 0,0 size 0x0
      on KeyDown: ActivateScreen("Alarm_Side", 0)

screen "Alarm_Side" 800x480
   AlarmView "Alarm view_1" at 0,0 size 799x426
   TextField "Text field_8" at 17,430 size 67x23; Text 'Prosess'
   TextField "Text field_9" at 125,430 size 53x23; Text 'Trend'
   TextField "Text field_10" at 225,430 size 52x23; Text 'Setup'
   TextField "Text field_16" at 29,450 size 40x23; Text 'Side'
   TextField "Text field_17" at 132,450 size 40x23; Text 'Side'
   TextField "Text field_18" at 230,450 size 40x23; Text 'Side'
   Softkey "Softkey_F1" at 0,0 size 0x0
      on KeyDown: ActivateScreen("Prosess_Side", 0)
   Softkey "Softkey_F2" at 0,0 size 0x0
      on KeyDown: ActivateScreen("Trend_Side", 0)
   Softkey "Softkey_F3" at 0,0 size 0x0
      on KeyDown: ActivateScreen("Setup_Side", 0)

screen "Trend_Side" 800x480
   TrendView "Trend view_1" at 170,0 size 630x430
   IOField "I/O field_1" at 70,110 size 90x40; FormatPattern s999.9
      ProcessValue <- "PID_Pump1_Control_sRet_r_Ctrl_Gain"
   IOField "I/O field_2" at 70,10 size 90x40; FormatPattern s999.9
      ProcessValue <- "HMI_LT_Level_SP"
   TextField "Text field_2" at 5,110 size 63x34; Text 'Gain'
   TextField "Text field_3" at 5,160 size 28x34; Text 'Ti'
   TextField "Text field_4" at 5,210 size 36x34; Text 'Td'
   IOField "I/O field_3" at 70,160 size 90x40; FormatPattern s999.9
      ProcessValue <- "PID_Pump1_Control_sRet_r_Ctrl_Ti"
   IOField "I/O field_4" at 70,210 size 90x40; FormatPattern s999.9
      ProcessValue <- "PID_Pump1_Control_sRet_r_Ctrl_Td"
   TextField "Text field_5" at 5,10 size 37x34; Text 'SP'
   IOField "I/O field_5" at 70,60 size 90x40; FormatPattern s999.9
      ProcessValue <- "DB_Equipment_LT01_Control_Sts_EU_Value_Out"
   TextField "Text field_6" at 5,60 size 38x34; Text 'PV'
   TextField "Text field_7" at 5,260 size 58x34; Text 'Man'
   TextField "Text field_8" at 24,430 size 52x23; Text 'Setup'
   TextField "Text field_9" at 117,430 size 67x23; Text 'Prosess'
   TextField "Text field_10" at 225,430 size 54x23; Text 'Alarm'
   TextField "Text field_16" at 29,450 size 40x23; Text 'Side'
   TextField "Text field_17" at 132,450 size 40x23; Text 'Side'
   TextField "Text field_18" at 230,450 size 40x23; Text 'Side'
   Switch "Switch_1" at 70,260 size 64x32; TextOn 'ON'; CaptionText 'Switch'; TextOff 'OFF'
      ProcessValue <- "DB_Equipment_Pumpe_01_Kontroll_Cmd_Auto_Start_Pumpe"
   Softkey "Softkey_F1" at 0,0 size 0x0
      on KeyDown: ActivateScreen("Setup_Side", 0)
   Softkey "Softkey_F2" at 0,0 size 0x0
      on KeyDown: ActivateScreen("Prosess_Side", 0)
   Softkey "Softkey_F3" at 0,0 size 0x0
      on KeyDown: ActivateScreen("Alarm_Side", 0)

screen "Setup_Side" 800x480
   TextField "Text field_1" at 230,5 size 329x43; Text 'Team Level Legends'
   IOField "I/O field_1" at 80,150 size 90x40; FormatPattern s999.9
      ProcessValue <- "PID_Pump1_Control_sRet_r_Ctrl_Gain"
   IOField "I/O field_2" at 80,50 size 90x40; FormatPattern s999.9
      ProcessValue <- "HMI_LT_Level_SP"
   TextField "Text field_2" at 10,150 size 63x34; Text 'Gain'
   TextField "Text field_3" at 10,200 size 28x34; Text 'Ti'
   TextField "Text field_4" at 10,250 size 36x34; Text 'Td'
   IOField "I/O field_3" at 80,200 size 90x40; FormatPattern s999.9
      ProcessValue <- "PID_Pump1_Control_sRet_r_Ctrl_Ti"
   IOField "I/O field_4" at 80,250 size 90x40; FormatPattern s999.9
      ProcessValue <- "PID_Pump1_Control_sRet_r_Ctrl_Td"
   TextField "Text field_5" at 10,50 size 37x34; Text 'SP'
   IOField "I/O field_5" at 80,100 size 90x40; FormatPattern s999.9
      ProcessValue <- "DB_Equipment_LT01_Control_Sts_EU_Value_Out"
   TextField "Text field_6" at 10,100 size 38x34; Text 'PV'
   TextField "Text field_7" at 370,170 size 335x34; Text 'Pumpe 01 Manuell kjøring'
   IOField "I/O field_7" at 690,50 size 90x40; FormatPattern s999.9
      ProcessValue <- "DB_Equipment_LT01_Control_Par_EU_Min"
   TextField "Text field_11" at 348,230 size 336x34; Text 'Manuelt Pådrag Pumpe 01'
   IOField "I/O field_9" at 694,230 size 90x40; FormatPattern s999.9
      ProcessValue <- "DB_Equipment_HMI_Control_Pump1_Par_HMI_Manual_Speed_Ref"
   TextField "Text field_12" at 505,50 size 166x34; Text 'LT 01 EU Min'
   IOField "I/O field_10" at 690,110 size 90x40; FormatPattern s999.9
      ProcessValue <- "DB_Equipment_LT01_Control_Par_EU_Max"
   TextField "Text field_13" at 505,110 size 172x34; Text 'LT 01 EU Max'
   TextField "Text field_14" at 10,300 size 200x34; Text 'Start Pumpe 01'
   TextField "Text field_15" at 10,380 size 211x34; Text 'Stopp Pumpe 01'
   Button "Button_4" at 230,300 size 96x32; TextOff 'Start'
      on Press: function_b14e0dd5("DB_Equipment_Pumpe_01_Kontroll_Cmd_Man_Start_Pumpe", 0)
   Button "Button_5" at 230,380 size 96x32; TextOff 'Stopp'
      on Press: function_b14e0dd5("DB_Equipment_Pumpe_01_Kontroll_Cmd_Man_Stop_Pumpe", 0)
   Switch "Switch_1" at 720,170 size 64x32; TextOn 'ON'; CaptionText 'Switch'; TextOff 'OFF'
      ProcessValue <- "DB_Equipment_Pumpe_01_Kontroll_Cmd_Auto_Start_Pumpe"
   TextField "Text field_8" at 17,430 size 67x23; Text 'Prosess'
   TextField "Text field_9" at 125,430 size 53x23; Text 'Trend'
   TextField "Text field_10" at 225,430 size 54x23; Text 'Alarm'
   TextField "Text field_16" at 29,450 size 40x23; Text 'Side'
   TextField "Text field_17" at 132,450 size 40x23; Text 'Side'
   TextField "Text field_18" at 230,450 size 40x23; Text 'Side'
   TextField "Text field_19" at 460,344 size 22x34; Text 'Text'
   TextField "Text field_20" at 332,300 size 353x34; Text 'Aktuell hastighet Pumpe 01'
   IOField "I/O field_6" at 694,300 size 90x40; FormatPattern s999.9
      ProcessValue <- "PID_Pumpe_01_Kontroll_Output"
   TextField "Text field_21" at 403,370 size 281x34; Text 'PID pådrag Pumpe 01'
   TextField "Text field_22" at 134,339 size 83x34; Text 'Kjører'
      Visibility <- "DI_P01_Run"
   Circle "Circle_1" at 262,341 size 32x32
      Appearance <- "DB_Equipment_Pumpe_01_Kontroll_Sts_Pumpe_Status"
   IOField "I/O field_8" at 694,370 size 90x40; FormatPattern s999.9
      ProcessValue <- "PID_Pumpe_01_Kontroll_Output"
   Softkey "Softkey_F1" at 0,0 size 0x0
      on KeyDown: ActivateScreen("Prosess_Side", 0)
   Softkey "Softkey_F2" at 0,0 size 0x0
      on KeyDown: ActivateScreen("Trend_Side", 0)
   Softkey "Softkey_F3" at 0,0 size 0x0
      on KeyDown: ActivateScreen("Alarm_Side", 0)
*)